FUNCTION "LKinCtrl_FwdFrame" : Void   // FC35005, SCL
TITLE = LKinCtrl_FwdFrame
{ S7_Optimized_Access := 'TRUE' }
AUTHOR : tech.team.motioncontrol@siemens.com
FAMILY : LKinCtrl
VERSION : 1.1
// Functionality: This function is calculating a forward frame transformation (-> In: Position in frame, Out: Position without frame)
// Support: tech.team.motioncontrol@siemens.com
// Note: Parameter comments are only available in language 'English (United States)'
   VAR_INPUT
      xIn : LReal;   // Input value x
      yIn : LReal;   // Input value y
      zIn : LReal;   // Input value z
      mode : Int;   // 0: Rotation + Translation, else: Rotation only
      frame : "LKinCtrl_typeFrame";   // Frame
   END_VAR
   VAR_OUTPUT
      xOut : LReal;   // Output value x
      yOut : LReal;   // Output value y
      zOut : LReal;   // Output value z
   END_VAR
   VAR_TEMP
      tempX1 : LReal;
      tempY1 : LReal;
      tempZ1 : LReal;
      tempX2 : LReal;
      tempY2 : LReal;
      tempZ2 : LReal;
      tempSin : LReal;
      tempCos : LReal;
   END_VAR
   // Ret_Val : Return value
   VAR CONSTANT
      DEGRAD : LReal := 0.0174532925199433;
   END_VAR
BEGIN
   //================================================================================
   // SIEMENS AG
   // (c)Copyright 2018 All Rights Reserved
   //--------------------------------------------------------------------------------
   // Library: LKinCtrl 
   // Tested with: S7-1516T-3 PN
   // Engineering: TIA Portal V15
   // Restrictions: -
   // Requirements: S7-1500/S7-1500T FW 2.5
   // Functionality: LKinCtrl_FwdFrame
   // This function is calculating a forward frame transformation
   //                (-> In: Position in frame, Out: Position without frame)
   // Support: tech.team.motioncontrol@siemens.com
   // Note: Parameter comments are only available in language 'English (United States)'
   //--------------------------------------------------------------------------------
   // Change log table:
   // Version  Date       Expert in charge Changes applied
   // 01.00.00 29.03.2018 SF               created
   // 01.01.00 03.09.2018 SF               bugfix
   //================================================================================

   REGION INPUT
     #tempX1 := #xIn;
     #tempY1 := #yIn;
     #tempZ1 := #zIn;
   END_REGION

   REGION ROTATION
     //first step: rotate c -> b -> a
     //----------------------------------------------------------------------------
     IF (#frame.c <> 0.0) THEN //x-rotation neccessary?
       #tempSin := SIN(#frame.c * #DEGRAD);
       #tempCos := COS(#frame.c * #DEGRAD);
       //rotate
       #tempX2 := #tempX1;
       #tempY2 := #tempY1 * #tempCos - #tempZ1 * #tempSin;
       #tempZ2 := #tempY1 * #tempSin + #tempZ1 * #tempCos;
       //store  
       #tempX1 := #tempX2;
       #tempY1 := #tempY2;
       #tempZ1 := #tempZ2;
     END_IF;

     IF (#frame.b <> 0.0) THEN //y-rotation neccessary?
       #tempSin := SIN(#frame.b * #DEGRAD);
       #tempCos := COS(#frame.b * #DEGRAD);
       //rotate
       #tempX2 := #tempX1 * #tempCos + #tempZ1 * #tempSin;
       #tempY2 := #tempY1;
       #tempZ2 := - #tempX1 * #tempSin + #tempZ1 * #tempCos;
       //store  
       #tempX1 := #tempX2;
       #tempY1 := #tempY2;
       #tempZ1 := #tempZ2;
     END_IF;

     IF (#frame.a <> 0.0) THEN //z-rotation neccessary?
       #tempSin := SIN(#frame.a * #DEGRAD);
       #tempCos := COS(#frame.a * #DEGRAD);
       //rotate
       #tempX2 := #tempX1 * #tempCos - #tempY1 * #tempSin;
       #tempY2 := #tempX1 * #tempSin + #tempY1 * #tempCos;
       #tempZ2 := #tempZ1;
       //store  
       #tempX1 := #tempX2;
       #tempY1 := #tempY2;
       #tempZ1 := #tempZ2;
     END_IF;
   END_REGION

   REGION TRANSLATION
     IF #mode = 0 THEN
       //second step: translation/ shifting X,Y,Z
       //-------------------------------------------------------------------------
       IF (#frame.x <> 0.0) THEN
         #tempX1 := #tempX1 + #frame.x;
       END_IF;
       IF (#frame.y <> 0.0) THEN
         #tempY1 := #tempY1 + #frame.y;
       END_IF;
       IF (#frame.z <> 0.0) THEN
         #tempZ1 := #tempZ1 + #frame.z;
       END_IF;
     END_IF;
   END_REGION

   REGION OUTPUT
     #xOut := #tempX1;
     #yOut := #tempY1;
     #zOut := #tempZ1;
   END_REGION
END_FUNCTION

FUNCTION "LKinCtrl_InvFrame" : Void   // FC35006, SCL
TITLE = LKinCtrl_InvFrame
{ S7_Optimized_Access := 'TRUE' }
AUTHOR : tech.team.motioncontrol@siemens.com
FAMILY : LKinCtrl
VERSION : 1.1
// Functionality: This function is calculating a inverse frame transformation (-> In: Position without frame, Out: Position in frame)
// Support: tech.team.motioncontrol@siemens.com
// Note: Parameter comments are only available in language 'English (United States)'
   VAR_INPUT
      xIn : LReal;   // Input value x
      yIn : LReal;   // Input value y
      zIn : LReal;   // Input value z
      mode : Int;   // 0: Rotation + Translation, else: Rotation only
      frame : "LKinCtrl_typeFrame";   // Frame
   END_VAR
   VAR_OUTPUT
      xOut : LReal;   // Output value x
      yOut : LReal;   // Output value y
      zOut : LReal;   // Output value z
   END_VAR
   VAR_TEMP
      tempX1 : LReal;
      tempY1 : LReal;
      tempZ1 : LReal;
      tempX2 : LReal;
      tempY2 : LReal;
      tempZ2 : LReal;
      tempSin : LReal;
      tempCos : LReal;
   END_VAR
   // Ret_Val : Return value
   VAR CONSTANT
      DEGRAD : LReal := 0.0174532925199433;
   END_VAR
BEGIN
   //================================================================================
   // SIEMENS AG
   // (c)Copyright 2018 All Rights Reserved
   //--------------------------------------------------------------------------------
   // Library: LKinCtrl
   // Tested with: S7-1516T-3 PN
   // Engineering: TIA Portal V15
   // Restrictions: -
   // Requirements: S7-1500/S7-1500T FW 2.5
   // Functionality: LKinCtrl_InvFrame
   // This function is calculating a inverse frame transformation
   //                (-> In: Position without frame, Out: Position in frame)
   // Support: tech.team.motioncontrol@siemens.com
   // Note: Parameter comments are only available in language 'English (United States)'
   //--------------------------------------------------------------------------------
   // Change log table:
   // Version  Date       Expert in charge Changes applied
   // 01.00.00 29.03.2018 SF               created
   // 01.01.00 03.09.2018 SF               bugfix
   //================================================================================

   REGION INPUT
     #tempX1 := #xIn;
     #tempY1 := #yIn;
     #tempZ1 := #zIn;
   END_REGION

   REGION TRANSLATION
     IF #mode = 0 THEN
       //first step: translation/ shifting X,Y,Z
       //-------------------------------------------------------------------------
       IF (#frame.x <> 0.0) THEN
         #tempX1 := #tempX1 - #frame.x;
       END_IF;
       IF (#frame.y <> 0.0) THEN
         #tempY1 := #tempY1 - #frame.y;
       END_IF;
       IF (#frame.z <> 0.0) THEN
         #tempZ1 := #tempZ1 - #frame.z;
       END_IF;
     END_IF;
   END_REGION

   REGION ROTATION
     //second step: rotate a -> b -> c
     //---------------------------------------------------------------------------
     IF (#frame.a <> 0.0) THEN //z-rotation neccessary?
       #tempSin := SIN(#frame.a * #DEGRAD);
       #tempCos := COS(#frame.a * #DEGRAD);
       //rotate
       #tempX2 := #tempX1 * #tempCos + #tempY1 * #tempSin;
       #tempY2 := - #tempX1 * #tempSin + #tempY1 * #tempCos;
       #tempZ2 := #tempZ1;
       //store  
       #tempX1 := #tempX2;
       #tempY1 := #tempY2;
       #tempZ1 := #tempZ2;
     END_IF;

     IF (#frame.b <> 0.0) THEN //y-rotation neccessary?
       #tempSin := SIN(#frame.b * #DEGRAD);
       #tempCos := COS(#frame.b * #DEGRAD);
       //rotate
       #tempX2 := #tempX1 * #tempCos - #tempZ1 * #tempSin;
       #tempY2 := #tempY1;
       #tempZ2 := #tempX1 * #tempSin + #tempZ1 * #tempCos;
       //store  
       #tempX1 := #tempX2;
       #tempY1 := #tempY2;
       #tempZ1 := #tempZ2;
     END_IF;

     IF (#frame.c <> 0.0) THEN //x-rotation neccessary?
       #tempSin := SIN(#frame.c * #DEGRAD);
       #tempCos := COS(#frame.c * #DEGRAD);
       //rotate
       #tempX2 := #tempX1;
       #tempY2 := #tempY1 * #tempCos + #tempZ1 * #tempSin;
       #tempZ2 := - #tempY1 * #tempSin + #tempZ1 * #tempCos;
       //store  
       #tempX1 := #tempX2;
       #tempY1 := #tempY2;
       #tempZ1 := #tempZ2;
     END_IF;
   END_REGION

   REGION OUTPUT
     #xOut := #tempX1;
     #yOut := #tempY1;
     #zOut := #tempZ1;
   END_REGION
END_FUNCTION

FUNCTION "LKinCtrl_FrameTrans" : Void   // FC35007, SCL
TITLE = LKinCtrl_FrameTrans
{ S7_Optimized_Access := 'TRUE' }
AUTHOR : tech.team.motioncontrol@siemens.com
FAMILY : LKinCtrl
VERSION : 2.0
// The FC calculates a given position transformed into or from another coordinate system depending on the actual / previous coordinate system of the cmd
   VAR_INPUT
      coordSystem : DInt;   // actual coordinate system
      coordSystemOld : DInt;   // previous coordinate system
      OCSFrames : Array[1..3] of "LKinCtrl_typeFrame";   // frame parameters read from TO_Kinematics
   END_VAR
   VAR_IN_OUT
      position : Array[1..4] of LReal;   // position to be transformed
   END_VAR
BEGIN
   //==========================================================================================
   // SIEMENS AG
   // (c)Copyright 2020 All Rights Reserved
   //------------------------------------------------------------------------------------------
   // Library: LKinCtrl
   // Tested with: S7-1517T-3 PN/DP
   // Engineering: TIA Portal V15
   // Restrictions: ---
   // Requirements: S7-1500T FW 2.5
   // Functionality: LKinCtrl_FrameTrans
   // The FC calculates a given position transformed into or from another coordinate system
   // depending on the actual / previous coordinate system of the cmd
   // 
   // Support: tech.team.motioncontrol@siemens.com
   // Note: Parameter comments are only available in language 'English (United States)'
   //------------------------------------------------------------------------------------------
   // Change log table:
   // Version    Date          Expert in charge    Changes applied
   // 01.00.00   16.04.2019    JR                  First release version v1.0
   // 02.00.00   14.04.2020    FR                  Use array of frames
   //===========================================================================================

   // Check if last CS differs from actual CS
   IF #coordSystem = #coordSystemOld THEN
     // No calculation needed --> Return
     RETURN;
   END_IF;

   // Calc new position
   // =================
   // Check if last CS was a OCS
   // YES: Transform position to WCS
   // NO: Do nothing --> Position is already in WCS
   IF (#coordSystemOld >= "CS_OCS1" AND #coordSystemOld <= "CS_OCS3") THEN
     // Get frame to WCS
     // foward frame transformation of lastPos to interprete position in WCS instead of OCS[1..3]
     "LKinCtrl_FwdFrame"(xIn := #position[1],
                         yIn := #position[2],
                         zIn := #position[3],
                         mode := 0,
                         frame := #OCSFrames[#coordSystemOld],
                         xOut => #position[1],
                         yOut => #position[2],
                         zOut => #position[3]);

     // Add "a" rotation to pos[4]
     // Rotation is needed because no change of orientation shall be done
     #position[4] := #position[4] + #OCSFrames[#coordSystemOld].a;
   ELSE
     ; // We are already in WCS
   END_IF;

   // Check if target CS is a OCS
   // YES: Transform position to target OCS
   // NO: Target CS is WCS --> Position is already in WCS from above
   IF (#coordSystem >= "CS_OCS1" AND #coordSystem <= "CS_OCS3") THEN
     // Get frame to target OCS
     // inverse frame transformation of lastPos to interprete position in OCS[1..3] instead of WCS
     "LKinCtrl_InvFrame"(xIn := #position[1],
                         yIn := #position[2],
                         zIn := #position[3],
                         mode := 0,
                         frame := #OCSFrames[#coordSystem],
                         xOut => #position[1],
                         yOut => #position[2],
                         zOut => #position[3]);

     // Substract "a" rotation to pos[4]
     // Rotation is needed because no change of orientation shall be done
     #position[4] := #position[4] - #OCSFrames[#coordSystem].a;
   ELSE
     ; // We are already in WCS
   END_IF;
END_FUNCTION

FUNCTION "LKinCtrl_ConvCircMode3To1" : Word   // FC35008, SCL
TITLE = LKinCtrl_ConvCircMode3To1
{ S7_Optimized_Access := 'TRUE' }
AUTHOR : tech.team.motioncontrol@siemens.com
FAMILY : LKinCtrl
VERSION : 2.0
// The FC converts a circular motion command programmed with circMode 3 (GCode) to a circular command programmed with circMode 1 (center point and arc given)
   VAR_INPUT
      coordinates : Variant;   // endPoint from path data element
      lastPos : Array[1..4] of LReal;   // previous last position
   END_VAR
   VAR_OUTPUT
      errorMessage : String;   // error message
   END_VAR
   VAR_IN_OUT
      cmdType : Int;   // cmdType of path data element
      circleParameters : "LKinCtrl_typeCircleParameters";   // circle parameters of path data element
   END_VAR
   VAR_TEMP
      tempAuxPoint : Array[1..3] of LReal;   // resulting auxPoint
      tempEndPointResult : Array[1..4] of LReal;   // resulting endPoint
      tempOM : Array[1..2] of LReal;   // temporary math variable
      tempMS : Array[1..2] of LReal;   // temporary math variable
      tempME : Array[1..2] of LReal;   // temporary math variable
      tempAxisVector : Array[1..2] of LReal;   // temporary math variable
      tempScalarProd_ME_Axis : LReal;   // temporary math variable
      tempScalarProd_MS_Axis : LReal;   // temporary math variable
      tempLength_ME : LReal;   // temporary math variable
      tempLength_MS : LReal;   // temporary math variable
      tempAngleME_rad : LReal;   // temporary math variable
      tempAngleMS_rad : LReal;   // temporary math variable
      tempAngleME_deg : LReal;   // temporary math variable
      tempAngleMS_deg : LReal;   // temporary math variable
      tempAngleDiff_deg : LReal;   // temporary math variable
      tempCtr : Int;   // temporary counter
      tempCoordinatesArray : REF_TO Array[1..4] of LReal;   // reference to coordinates from pre buf element
      tempCoordinatesStruct : REF_TO "LKinCtrl_typeCartesianPosition";   // reference to coordinates from normal element
      tempCoordinates : Array[1..4] of LReal;   // temporary array for input end point
   END_VAR
   // Ret_Val : return value
   VAR CONSTANT
      ERR_INVALID_CMDTYPE : Word := 16#8265;   // error due to invalid cmdType
      STATUS_NO_ERROR : Word := 16#0;   // status no error occured
   END_VAR
BEGIN
   //==========================================================================================
   // SIEMENS AG
   // (c)Copyright 2020 All Rights Reserved
   //------------------------------------------------------------------------------------------
   // Library: LKinCtrl
   // Tested with: S7-1517T-3 PN/DP
   // Engineering: TIA Portal V15
   // Restrictions: ---
   // Requirements: S7-1500T FW 2.5
   // Functionality: LKinCtrl_ConvCircMode3To1
   // The FC converts a circular motion command programmed with circMode 3 (GCode) to a circular
   // command programmed with circMode 1 (center point and arc given)
   // 
   // Support: tech.team.motioncontrol@siemens.com
   // Note: Parameter comments are only available in language 'English (United States)'
   //------------------------------------------------------------------------------------------
   // Change log table:
   // Version    Date          Expert in charge    Changes applied
   // 01.00.00   03.07.2019    JR                  First release version v1.0
   // 02.00.00   06.04.2020    FR                  Changed interface to fit PathDataPreBuf and normal element
   //===========================================================================================

   IF TypeOf(#coordinates) = LKinCtrl_typeCartesianPosition THEN
     // Assignment
     #tempCoordinatesStruct ?= #coordinates;

     // Assign temp with values
     #tempCoordinates[1] := #tempCoordinatesStruct<?OpDeref?>.x;
     #tempCoordinates[2] := #tempCoordinatesStruct<?OpDeref?>.y;
     #tempCoordinates[3] := #tempCoordinatesStruct<?OpDeref?>.z;
     #tempCoordinates[4] := #tempCoordinatesStruct<?OpDeref?>.a;

   ELSIF TypeOfElements(#coordinates) = LReal AND IS_ARRAY(#coordinates) AND CountOfElements(#coordinates) = 4 THEN
     // Assignment
     #tempCoordinatesArray ?= #coordinates;

     // Assign temp with values
     #tempCoordinates := #tempCoordinatesArray<?OpDeref?>;

   ELSE
     ; // Wrong input ?
   END_IF;

   // add conversion of circMode CM: 3 circular cmds -> CM: 1
   IF (#cmdType = "LKINCTRL_MC_MOVECIRCULARABS"
     OR #cmdType = "LKINCTRL_MC_MOVECIRCULARREL")
     AND #circleParameters.circMode = 3
   THEN

     // conversion relative to absoulte for auxPoint (and EndPoint)
     FOR #tempCtr := 1 TO 3 DO
       // always convert auxPoint ==> always relative in this circle definition
       // add new auxPoint as incremental value to last position
       #tempAuxPoint[#tempCtr] := #lastPos[#tempCtr] + #circleParameters.auxPoint[#tempCtr];
       // copy edited auxPoint to command for later use
       #circleParameters.auxPoint[#tempCtr] := #tempAuxPoint[#tempCtr];
     END_FOR;

     // only convert endPoint in case of relative command
     IF #cmdType = "LKINCTRL_MC_MOVECIRCULARREL" THEN
       #tempEndPointResult[1] := #lastPos[1] + #tempCoordinates[1];
       #tempEndPointResult[2] := #lastPos[2] + #tempCoordinates[2];
       #tempEndPointResult[3] := #lastPos[3] + #tempCoordinates[3];
       #tempEndPointResult[4] := #lastPos[4] + #tempCoordinates[4];
       #cmdType := "LKINCTRL_MC_MOVECIRCULARABS";
     ELSE
       #tempEndPointResult := #tempCoordinates;
     END_IF;

     // change circMode = 3 (define center and endPoint) to circMode = 1 (define center and arc)
     #circleParameters.circMode := 1;

     // different behavior for different circlePlanes - write input vectors to calc variables 2D
     // 0: ciclePlane XZ
     IF #circleParameters.circlePlane = 0 THEN

       // vector origin to circle center point 
       #tempOM[1] := #tempAuxPoint[1];
       #tempOM[2] := #tempAuxPoint[3];

       // unit vector x axis
       #tempAxisVector[1] := 1;
       #tempAxisVector[2] := 0;

       // vector circle center point to start point
       #tempMS[1] := #lastPos[1] - #tempOM[1];
       #tempMS[2] := #tempOM[2] - #lastPos[3];

       // vector circle center point to end point
       #tempME[1] := #tempEndPointResult[1] - #tempOM[1];
       #tempME[2] := #tempOM[2] - #tempEndPointResult[3];

       // 1: ciclePlane YZ
     ELSIF #circleParameters.circlePlane = 1 THEN

       // vector origin to circle center point 
       #tempOM[1] := #tempAuxPoint[2];
       #tempOM[2] := #tempAuxPoint[3];

       // unit vector x axis ==> simulating y axis here due to moved commands
       #tempAxisVector[1] := 1;
       #tempAxisVector[2] := 0;

       // vector circle center point to start point
       #tempMS[1] := #lastPos[2] - #tempOM[1];
       #tempMS[2] := #lastPos[3] - #tempOM[2];

       // vector circle center point to end point
       #tempME[1] := #tempEndPointResult[2] - #tempOM[1];
       #tempME[2] := #tempEndPointResult[3] - #tempOM[2];

       // 2: ciclePlane XY
     ELSIF #circleParameters.circlePlane = 2 THEN

       // vector origin to circle center point 
       #tempOM[1] := #tempAuxPoint[1];
       #tempOM[2] := #tempAuxPoint[2];

       // unit vector x axis
       #tempAxisVector[1] := 1;
       #tempAxisVector[2] := 0;


       // vector circle center point to start point
       #tempMS[1] := #lastPos[1] - #tempOM[1];
       #tempMS[2] := #lastPos[2] - #tempOM[2];

       // vector circle center point to end point
       #tempME[1] := #tempEndPointResult[1] - #tempOM[1];
       #tempME[2] := #tempEndPointResult[2] - #tempOM[2];

     ELSE
       // error ==> wrong circlePlane
       ;
     END_IF;

     // VECTOR CALCULATIONS
     // calc scalar product of ME (circle center point to end point) with x axis
     #tempScalarProd_ME_Axis := "LKinCtrl_VecScalarProd_2D"(vIn1 := #tempME, vIn2 := #tempAxisVector);
     // calc scalar product of MS (circle center point to start point / LastPos) with x axis
     #tempScalarProd_MS_Axis := "LKinCtrl_VecScalarProd_2D"(vIn1 := #tempMS, vIn2 := #tempAxisVector);

     // calc vector length ME
     #tempLength_ME := "LKinCtrl_VecAbs_2D"(#tempME);
     // calc vector length MS
     #tempLength_MS := "LKinCtrl_VecAbs_2D"(#tempMS);

     // calc angle ME to axis
     #tempAngleME_rad := ACOS(#tempScalarProd_ME_Axis / (#tempLength_ME * 1));

     IF #tempME[2] <= 0 THEN
       // invert angle due to ACOS range (only 0..PI)
       #tempAngleME_rad := 2 * "LKINCTRL_PI" - #tempAngleME_rad;
     ELSE
       ;
     END_IF;
     // convert to degrees
     #tempAngleME_deg := #tempAngleME_rad * 180 / "LKINCTRL_PI";

     // calc angle MS to axis
     #tempAngleMS_rad := ACOS(#tempScalarProd_MS_Axis / (#tempLength_MS * 1));
     // check for vector Ms to point downwards (below ! (x) axis)
     IF #tempMS[2] < 0 THEN
       // invert angle due to ACOS range
       #tempAngleMS_rad := 2 * "LKINCTRL_PI" - #tempAngleMS_rad;
     ELSE
       ;
     END_IF;
     // convert to degrees
     #tempAngleMS_deg := #tempAngleMS_rad * 180 / "LKINCTRL_PI";


     // separation of path choice for angle calculation
     // 0: CCW - counterclockwise / mathematical positive angle
     IF #circleParameters.pathChoice = 0 THEN
       // calculate difference angle
       #tempAngleDiff_deg := #tempAngleME_deg - #tempAngleMS_deg;
       IF #tempAngleDiff_deg > 0 THEN
         // write caclulated angle
         #circleParameters.arc := #tempAngleDiff_deg;
       ELSE
         // write caclulated angle ==> add 360 degrees to get positive angle value
         #circleParameters.arc := #tempAngleDiff_deg + 360;
       END_IF;

       // 1: CW - clockwise / mathematical negative angle
     ELSIF #circleParameters.pathChoice = 1 THEN
       // calculate difference angle
       #tempAngleDiff_deg := #tempAngleMS_deg - #tempAngleME_deg;
       IF #tempAngleDiff_deg >(* = *) 0 THEN
         // write caclulated angle
         #circleParameters.arc := #tempAngleDiff_deg;
       ELSE
         // write caclulated angle ==> add 360 degrees to get positive angle value
         #circleParameters.arc := #tempAngleDiff_deg + 360;
       END_IF;

     ELSE
       // wrong input for pathChoice
       ;
     END_IF;
     // conversion successful
     #LKinCtrl_ConvCircMode3To1 := #STATUS_NO_ERROR;

   ELSE
     // do nothing
     #LKinCtrl_ConvCircMode3To1 := #ERR_INVALID_CMDTYPE;
     #errorMessage := 'no circular command to convert';
   END_IF;
END_FUNCTION

FUNCTION "LKinCtrl_EvaluateParamValidBits" : Void   // FC35009, SCL
TITLE = LKinCtrl_EvaluateParamValidBits
{ S7_Optimized_Access := 'TRUE' }
AUTHOR : tech.team.motioncontrol@siemens.com
FAMILY : LKinCtrl
VERSION : 1.0
// The FC evaluates the parameterValid bits of a given command and copies the coordinates for valid bits and overwrites coordinates by last position or 0.0 increment for invalid bits.
   VAR_INPUT
      parameterValidBits : Array[1.."LKINCTRL_NO_OF_VALID_BITS"] of Bool;   // parameter valid bits of actual command
      lastPos : Array[1..4] of LReal;   // previous last position
   END_VAR
   VAR_OUTPUT
      errorMessage : String;   // error message
   END_VAR
   VAR_IN_OUT
      command : "LKinCtrl_typePathDataElement";   // command to evaluate and edit
   END_VAR
   VAR_TEMP
      tempPosElemCtr : Int;   // temporary counter variable
   END_VAR
BEGIN
   //==========================================================================================
   // SIEMENS AG
   // (c)Copyright 2019 All Rights Reserved
   //------------------------------------------------------------------------------------------
   // Library: LKinCtrl
   // Tested with: S7-1517T-3 PN/DP
   // Engineering: TIA Portal V15
   // Restrictions: ---
   // Requirements: S7-1500T FW 2.5
   // Functionality: LKinCtrl_EvaluateParamValidBits
   // The FC evaluates the parameterValid bits of a given command and copies the coordinates for
   // valid bits and overwrites coordinates by last position or 0.0 increment for invalid bits.
   // 
   // Support: tech.team.motioncontrol@siemens.com
   // Note: Parameter comments are only available in language 'English (United States)'
   //------------------------------------------------------------------------------------------
   // Change log table:
   // Version    Date          Expert in charge    Changes applied
   // 01.00.00   08.07.2019    JR                  First release version v1.0
   // 01.00.01   09.08.2019    JR                  excluded auxPoint from parameter valid bits
   //===========================================================================================

   // ParameterValid bit check
   //====================================================================================================================================

   // -----------------------------------------------------------------------------------
   IF #command.cmdType = "LKINCTRL_MC_MOVELINEARABS" OR #command.cmdType = "LKINCTRL_MC_MOVECIRCULARABS" THEN

     FOR #tempPosElemCtr := 1 TO "LKINCTRL_NO_OF_VALID_BITS" DO
       // Check valid bits and copy last pos (X,Y,Z,A) where missing
       IF #parameterValidBits[#tempPosElemCtr] = FALSE THEN
         // write lastPos as target pos if invalid
         IF #tempPosElemCtr = 1 THEN
           #command.cmdCoordinates.cartesianPosition.x := #lastPos[#tempPosElemCtr];
         ELSIF #tempPosElemCtr = 2 THEN
           #command.cmdCoordinates.cartesianPosition.y := #lastPos[#tempPosElemCtr];
         ELSIF #tempPosElemCtr = 3 THEN
           #command.cmdCoordinates.cartesianPosition.z := #lastPos[#tempPosElemCtr];
         ELSIF #tempPosElemCtr = 4 THEN
           #command.cmdCoordinates.cartesianPosition.a := #lastPos[#tempPosElemCtr];
         END_IF;

         // // exclude auxPoint from parameterValidBits, add additional parameterValidBits if needed
         // // write lastPos to auxPoint if invalid
         // IF #tempPosElemCtr < 4 THEN
         //   #command.cmdParameters.circleParameters.auxPoint[#tempPosElemCtr] := #lastPos[#tempPosElemCtr];
         // ELSE
         //   ; // do not copy for tempPosElemCtr = 4
         // END_IF;
       ELSE
         ; // Keep programmed position from #pathDataElementPreBuf.cmdCoordinates.cartesianPosition
       END_IF;
     END_FOR;

   ELSIF #command.cmdType = "LKINCTRL_MC_MOVELINEARREL" OR #command.cmdType = "LKINCTRL_MC_MOVECIRCULARREL" THEN
     FOR #tempPosElemCtr := 1 TO "LKINCTRL_NO_OF_VALID_BITS" DO
       // Check valid bits and set absolute pos to 0.0 (X,Y,Z,A)
       IF #parameterValidBits[#tempPosElemCtr] = FALSE THEN
         // write no increment as relative target pos if invalid
         IF #tempPosElemCtr = 1 THEN
           #command.cmdCoordinates.cartesianPosition.x := 0.0;
         ELSIF #tempPosElemCtr = 2 THEN
           #command.cmdCoordinates.cartesianPosition.y := 0.0;
         ELSIF #tempPosElemCtr = 3 THEN
           #command.cmdCoordinates.cartesianPosition.z := 0.0;
         ELSIF #tempPosElemCtr = 4 THEN
           #command.cmdCoordinates.cartesianPosition.a := 0.0;
         END_IF;

         // // exclude auxPoint from parameterValidBits, add additional parameterValidBits if needed
         // // write no increment as relative target pos if invalid
         // IF #tempPosElemCtr < 4 THEN
         //   #command.cmdParameters.circleParameters.auxPoint[#tempPosElemCtr] := 0.0;
         // ELSE
         //   ; // do not copy for tempPosElemCtr = 4
         // END_IF;
       ELSE
         ; // Keep programmed position from #pathDataElementPreBuf.cmdCoordinates.cartesianPosition
       END_IF;
     END_FOR;
   ELSE
     ; // Nothing to do for this cmdType
   END_IF;
END_FUNCTION

FUNCTION "LKinCtrl_CallMC_TrackConv_PosAxis" : Void   // FC35010, SCL
TITLE = LKinCtrl_CallMC_TrackConv_PosAxis
{ S7_Optimized_Access := 'TRUE' }
AUTHOR : tech.team.motioncontrol@siemens.com
FAMILY : LKinCtrl
VERSION : 1.0
// Call given MC_TrackConveyorBelt instance
   VAR_INPUT
      posAxis : TO_PositioningAxis;   // Positioning axis input
      axesGroup : TO_Kinematics;   // Kinematics input
   END_VAR
   VAR_IN_OUT
      instTrackConveyorBelt : MC_TRACKCONVEYORBELT;   // Instance of MC_TrackConveyorBelt to be called
   END_VAR
BEGIN
   //================================================================================
   // SIEMENS AG
   // (c)Copyright 2020 All Rights Reserved
   //--------------------------------------------------------------------------------
   // Library: LKinCtrl
   // Tested with: S7-1517T-3 PN
   // Engineering: TIA Portal V16
   // Restrictions: -
   // Requirements: S7-1500T FW 2.8
   // Functionality: Call MC_TrackConveyorBelt
   // Support: tech.team.motioncontrol@siemens.com
   // Note: Parameter comments are only available in language 'English (United States)'
   //-----------------------------------------------------------------------------
   // Change log table:
   // Version    Date          Expert in charge    Changes applied
   // 01.00.00   24.04.2020    FR                  First released version
   //===========================================================================================

   // call MC_TrackConveyorBelt
   #instTrackConveyorBelt(AxesGroup:=#axesGroup,
                              ConveyorBelt:=#posAxis);
END_FUNCTION

FUNCTION "LKinCtrl_CallMC_TrackConv_SyncAxis" : Void   // FC35011, SCL
TITLE = LKinCtrl_CallMC_TrackConv_SyncAxis
{ S7_Optimized_Access := 'TRUE' }
AUTHOR : tech.team.motioncontrol@siemens.com
FAMILY : LKinCtrl
VERSION : 1.0
// Call given MC_TrackConveyorBelt instance
   VAR_INPUT
      syncAxis : TO_SynchronousAxis;   // Synchronous axis input
      axesGroup : TO_Kinematics;   // Kinematics input
   END_VAR
   VAR_IN_OUT
      instTrackConveyorBelt : MC_TRACKCONVEYORBELT;   // Instance of MC_TrackConveyorBelt to be called
   END_VAR
BEGIN
   //================================================================================
   // SIEMENS AG
   // (c)Copyright 2020 All Rights Reserved
   //--------------------------------------------------------------------------------
   // Library: LKinCtrl
   // Tested with: S7-1517T-3 PN
   // Engineering: TIA Portal V16
   // Restrictions: -
   // Requirements: S7-1500T FW 2.8
   // Functionality: Call MC_TrackConveyorBelt
   // Support: tech.team.motioncontrol@siemens.com
   // Note: Parameter comments are only available in language 'English (United States)'
   //-----------------------------------------------------------------------------
   // Change log table:
   // Version    Date          Expert in charge    Changes applied
   // 01.00.00   24.04.2020    FR                  First released version
   //===========================================================================================

   // call MC_TrackConveyorBelt
   #instTrackConveyorBelt(AxesGroup := #axesGroup,
                          ConveyorBelt := #syncAxis);
END_FUNCTION

FUNCTION "LKinCtrl_CallMC_TrackConv_ExtEncoder" : Void   // FC35012, SCL
TITLE = LKinCtrl_CallMC_TrackConv_ExtEncoder
{ S7_Optimized_Access := 'TRUE' }
AUTHOR : tech.team.motioncontrol@siemens.com
FAMILY : LKinCtrl
VERSION : 1.0
// Call given MC_TrackConveyorBelt instance
   VAR_INPUT
      extEncoder : TO_ExternalEncoder;   // External Encoder input
      axesGroup : TO_Kinematics;   // Kinematics input
   END_VAR
   VAR_IN_OUT
      instTrackConveyorBelt : MC_TRACKCONVEYORBELT;   // Instance of MC_TrackConveyorBelt to be called
   END_VAR
BEGIN
   //================================================================================
   // SIEMENS AG
   // (c)Copyright 2020 All Rights Reserved
   //--------------------------------------------------------------------------------
   // Library: LKinCtrl
   // Tested with: S7-1517T-3 PN
   // Engineering: TIA Portal V16
   // Restrictions: -
   // Requirements: S7-1500T FW 2.8
   // Functionality: Call MC_TrackConveyorBelt
   // Support: tech.team.motioncontrol@siemens.com
   // Note: Parameter comments are only available in language 'English (United States)'
   //-----------------------------------------------------------------------------
   // Change log table:
   // Version    Date          Expert in charge    Changes applied
   // 01.00.00   24.04.2020    FR                  First released version
   //===========================================================================================

   // call MC_TrackConveyorBelt
   #instTrackConveyorBelt(AxesGroup := #axesGroup,
                          ConveyorBelt := #extEncoder);
END_FUNCTION

FUNCTION "LKinCtrl_CallMC_TrackConv_LeadingAxisProxy" : Void   // FC35013, SCL
TITLE = LKinCtrl_CallMC_TrackConv_LeadingAxisProxy
{ S7_Optimized_Access := 'TRUE' }
AUTHOR : tech.team.motioncontrol@siemens.com
FAMILY : LKinCtrl
VERSION : 1.0
// Call given MC_TrackConveyorBelt instance
   VAR_INPUT
      leadingAxisProxy : TO_LeadingAxisProxy;   // Leading axis proxy input
      axesGroup : TO_Kinematics;   // Kinematics input
   END_VAR
   VAR_IN_OUT
      instTrackConveyorBelt : MC_TRACKCONVEYORBELT;   // Instance of MC_TrackConveyorBelt to be called
   END_VAR
BEGIN
   //================================================================================
   // SIEMENS AG
   // (c)Copyright 2020 All Rights Reserved
   //--------------------------------------------------------------------------------
   // Library: LKinCtrl
   // Tested with: S7-1517T-3 PN
   // Engineering: TIA Portal V16
   // Restrictions: -
   // Requirements: S7-1500T FW 2.8
   // Functionality: Call MC_TrackConveyorBelt
   // Support: tech.team.motioncontrol@siemens.com
   // Note: Parameter comments are only available in language 'English (United States)'
   //-----------------------------------------------------------------------------
   // Change log table:
   // Version    Date          Expert in charge    Changes applied
   // 01.00.00   24.04.2020    FR                  First released version
   //===========================================================================================

   // call MC_TrackConveyorBelt
   #instTrackConveyorBelt(AxesGroup := #axesGroup,
                          ConveyorBelt := #leadingAxisProxy);
END_FUNCTION

FUNCTION "LKinCtrl_VecAbs_2D" : LReal   // FC35029, SCL
TITLE = LKinCtrl_VecAbs_2D
{ S7_Optimized_Access := 'TRUE' }
AUTHOR : tech.team.motioncontrol@siemens.com
FAMILY : LKinCtrl
VERSION : 1.0
// Calculates the length of a given vector in 2D
   VAR_INPUT
      vIn : Array[1..2] of LReal;   // Input vector
   END_VAR
   // Ret_Val : Output scalar
BEGIN
   //=============================================================================
   // SIEMENS AG
   // (c)Copyright 2019 All Rights Reserved
   //-----------------------------------------------------------------------------
   // Library: - 
   // Tested with: S7-1516T-3 PN
   // Engineering: TIA Portal V15
   // Restrictions: -
   // Requirements: S7-1500/S7-1500T FW 2.5
   // Functionality: Calculate length of vector
   //-----------------------------------------------------------------------------
   // Change log table:
   // Version  Date       Expert in charge Changes applied
   // 01.00.00 27.08.2018 SF               created
   // 01.00.01 29.01.2019 JR               adaptions for LKinCtrl 
   //=============================================================================

   #LKinCtrl_VecAbs_2D := SQRT((* #vIn[0]*#vIn[0] + *)#vIn[1]*#vIn[1] + #vIn[2]*#vIn[2]);
END_FUNCTION

FUNCTION "LKinCtrl_VecScalarProd_2D" : LReal   // FC35030, SCL
TITLE = LKinCtrl_VecScalarProd_2D / LKinCtrl_VecScalarProd
{ S7_Optimized_Access := 'TRUE' }
AUTHOR : tech.team.motioncontrol@siemens.com
FAMILY : LKinCtrl
VERSION : 1.0
// Calculates the scalar product of given vectors
   VAR_INPUT
      vIn1 : Array[1..2] of LReal;   // Input vector 1
      vIn2 : Array[1..2] of LReal;   // Input vector 2
   END_VAR
   // Ret_Val : Output scalar
BEGIN
   //=============================================================================
   // SIEMENS AG
   // (c)Copyright 2019 All Rights Reserved
   //-----------------------------------------------------------------------------
   // Library: - 
   // Tested with: S7-1516T-3 PN
   // Engineering: TIA Portal V15
   // Restrictions: -
   // Requirements: S7-1500/S7-1500T FW 2.5
   // Functionality: Scalar product of two coordinates
   //-----------------------------------------------------------------------------
   // Change log table:
   // Version  Date       Expert in charge Changes applied
   // 01.00.00 27.08.2018 SF               created
   // 01.00.01 29.01.2019 JR               adaptions for LKinCtrl 
   //=============================================================================

   #LKinCtrl_VecScalarProd_2D := (* #vIn1[0]*#vIn2[0] + *)#vIn1[1]*#vIn2[1] + #vIn1[2]*#vIn2[2];
END_FUNCTION

FUNCTION "LKinCtrl_GetPathDataCmd" : Word   // FC35031, SCL
TITLE = LKinCtrl_GetPathDataCmd
{ S7_Optimized_Access := 'TRUE' }
AUTHOR : tech.team.motioncontrol@siemens.com
FAMILY : LKinCtrl
VERSION : 1.0
// Copy the path command from any path data type at the given index
   VAR_INPUT
      pathDataType : USInt;   // Type of path data which is connected
      index : DInt;   // Index to be copied
      pathDataReduced : REF_TO "LKinCtrl_typePathData_reduced";   // Reference to reduced path data
      pathData : REF_TO "LKinCtrl_typePathData";   // Reference to normal path data
      pathDataAdvanced : REF_TO "LKinCtrl_typePathData_advanced";   // Reference to advanced path data
   END_VAR
   VAR_OUTPUT
      pathDataCommand : "LKinCtrl_typePathDataElement";   // Resulting path data command
      parameterValid : Array[1.."LKINCTRL_NO_OF_VALID_BITS"] of Bool;   // Resulting parameter valid bits
   END_VAR
   VAR_TEMP
      tempCtr : Int;   // Temporary counter
   END_VAR
   // Ret_Val : Return value
BEGIN
   //==========================================================================================
   // SIEMENS AG
   // (c)Copyright 2020 All Rights Reserved
   //------------------------------------------------------------------------------------------
   // Library: LKinCtrl
   // Tested with: S7-1517T-3 PN/DP
   // Engineering: TIA Portal V15
   // Restrictions: ---
   // Requirements: S7-1500T FW 2.5
   // Functionality: LKinCtrl_GetPathDataCmd
   // The FC copies the path data command at the given index to the output.
   // 
   // Support: tech.team.motioncontrol@siemens.com
   // Note: Parameter comments are only available in language 'English (United States)'
   //------------------------------------------------------------------------------------------
   // Change log table:
   // Version    Date          Expert in charge    Changes applied
   // 01.00.00   07.04.2020    FR                  First release version v1.0
   //===========================================================================================

   // Set return value
   #LKinCtrl_GetPathDataCmd := 16#00;

   // Copy actual path data element where index is pointing at
   IF #pathDataType = "LKINCTRL_PATHDATA_TYPE_REDUCED" THEN
     // Copy command
     #pathDataCommand.cmdType := #pathDataReduced<?OpDeref?>.commands[#index].cmdType;
     #pathDataCommand.cmdName := #pathDataReduced<?OpDeref?>.commands[#index].cmdName;
     #pathDataCommand.cmdActivated := #pathDataReduced<?OpDeref?>.commands[#index].cmdActivated; // !
     #pathDataCommand.cmdCoordinates := #pathDataReduced<?OpDeref?>.commands[#index].cmdCoordinates;
     #pathDataCommand.cmdParameters.pathDynamics := #pathDataReduced<?OpDeref?>.commands[#index].cmdParameters.pathDynamics;
     #pathDataCommand.cmdParameters.orientationDirection := #pathDataReduced<?OpDeref?>.commands[#index].cmdParameters.orientationDirection;
     #pathDataCommand.cmdParameters.bufferMode := #pathDataReduced<?OpDeref?>.commands[#index].cmdParameters.bufferMode;
     #pathDataCommand.cmdParameters.transitionParameters := #pathDataReduced<?OpDeref?>.commands[#index].cmdParameters.transitionParameters;
     #pathDataCommand.cmdParameters.dynamicAdaption := #pathDataReduced<?OpDeref?>.commands[#index].cmdParameters.dynamicAdaption;
     #pathDataCommand.setFlags := #pathDataReduced<?OpDeref?>.commands[#index].setFlags;
     #pathDataCommand.valueFlags := #pathDataReduced<?OpDeref?>.commands[#index].valueFlags;

     // always set valid bits to true
     FOR #tempCtr := 1 TO "LKINCTRL_NO_OF_VALID_BITS" DO
       // Statement section FOR
       #parameterValid[#tempCtr] := TRUE;
     END_FOR;

   ELSIF #pathDataType = "LKINCTRL_PATHDATA_TYPE_NORMAL" THEN
     // Copy command
     #pathDataCommand := #pathData<?OpDeref?>.commands[#index];

     // always set valid bits to true
     FOR #tempCtr := 1 TO "LKINCTRL_NO_OF_VALID_BITS" DO
       // Statement section FOR
       #parameterValid[#tempCtr] := TRUE;
     END_FOR;

   ELSIF #pathDataType = "LKINCTRL_PATHDATA_TYPE_ADVANCED" THEN
     // Copy command
     #pathDataCommand.cmdType := #pathDataAdvanced<?OpDeref?>.commands[#index].cmdType;
     #pathDataCommand.cmdName := #pathDataAdvanced<?OpDeref?>.commands[#index].cmdName;
     #pathDataCommand.cmdActivated := #pathDataAdvanced<?OpDeref?>.commands[#index].cmdActivated;
     #pathDataCommand.cmdCoordinates := #pathDataAdvanced<?OpDeref?>.commands[#index].cmdCoordinates;
     #pathDataCommand.cmdParameters := #pathDataAdvanced<?OpDeref?>.commands[#index].cmdParameters;
     #pathDataCommand.setFlags := #pathDataAdvanced<?OpDeref?>.commands[#index].setFlags;
     #pathDataCommand.valueFlags := #pathDataAdvanced<?OpDeref?>.commands[#index].valueFlags;

     // Copy valid bits from command
     #parameterValid := #pathDataAdvanced<?OpDeref?>.commands[#index].parameterValid;

   ELSE
     // Set return value to error
     #LKinCtrl_GetPathDataCmd := 16#01;
   END_IF;
END_FUNCTION

// folder: LKinLang_Blocks

FUNCTION_BLOCK "LKinLang_Parser"   // FB35450, SCL
TITLE = LKinLang_Parser
{ S7_Optimized_Access := 'TRUE' }
AUTHOR : tech.team.motioncontrol@siemens.com
FAMILY : LKinLang
VERSION : 1.3
// The FB parses strings from line buffer to PathData commands using different language
// packages.
// The FB parses strings from line buffer to PathData commands using different languagepackages.
   VAR_INPUT
      execute : Bool;   // Rising edge starts action once
      stop : Bool;   // Rising edge stops execution
      language : Int;   // Selected language to be parsed
      syntaxCheck : USInt;   // 0: No check before; 1: Check only; 2: Check and execute
      flagModeDefaults : "LKinLang_typeFlagModeDefaults";   // Structure to define default flag settings for setFlags and valueFlags
   END_VAR
   VAR_OUTPUT
      done : Bool;   // TRUE: Commanded functionality has been completed successfully
      busy : Bool;   // TRUE: FB is not finished and new output values can be expected
      commandAborted : Bool;   // TRUE: Commanded functionality has been aborted by another command
      error : Bool;   // TRUE: An error occurred during the execution of the FB
      status : Word := 16#7000;   // 16#0000 - 16#7FFF: Status of the FB, 16#8000 - 16#FFFF: Error identification
      errorString : String;   // Error description as string
   END_VAR
   VAR_IN_OUT
      lineBuffer : "LKinLang_typeLineBuffer";   // String buffer connection
      pathData : "LKinCtrl_typePathData_advanced";   // PathData connection
      preProcessConfig : "LKinLang_typePreProcessorReplacement";   // Array which defines replacements
      parameterDefaults : Variant;   // Structure to define default values in language (e.g. velocity for rapid linear)
      interfaceVariables : "LKinLang_typeInterfaceVariables";   // Interface variables arrays
   END_VAR
   VAR
      statExecuteOld : Bool;   // Old value of 'execute' input for edge detection
      statDone : Bool;   // Static value for output 'done'
      statBusy : Bool;   // Static value for output 'busy'
      statCommandAborted : Bool;   // Static value for output 'commandAborted'
      statError : Bool;   // Static value for output 'error'
      statStatus : Word := 16#7000;   // Static value for output 'status'
      statErrorString : String;   // Error string variable
      statStopOld : Bool;   // Static storing for the stop input
      statFBState : DInt := 0;   // State in the state machine of the FB
      statStateIntern : Int;   // Internal state variable
      statSelectedLanguage : Int;   // Selected Language
      statPositioningMode : Int := 1;   // Positioning mode: 1=Absolute, 2=Relative
      statPositioningModeOld : Int := 1;   // Last Positioning mode
      statLastIndexLookUp : DInt;   // Last found command in Language Package
      statLastIndexOfMerger : Int;   // Last entry in merger array
      statLookUpTableCounter : Int;   // Counter to continue look up table
      statAddPointer : Int;   // Internal static to for the PathData add pointer
      statActualValueFlagNumber : Int;   // Static storing for the actual value flag number
      statActualFlagNumber : Int;   // Static storing for the actual boolean flag number
      statStringExpression : String;   // Static storing for the string expression
      statRightSideOfEquation : Bool;   // Static storing if right side of equation
      statDirectCmdWord : Word;   // Static storing direct command word
      statSyntaxCheck : USInt;   // Static storing for syntaxCheck input
      statSearchedLine : UDInt;   // Static storing for requested line number
      statConfigCmdWords : Array[1.."LKINLANG_NUMBER_OF_FOLLOW_VALUES"] of Word;   // Static storing config command word
      statTokenCheck : Struct   // Static struct with the token to check
         actual : String;
         previous : String;
      END_STRUCT;
      statTokenizedLine : "LKinLang_typeLineTokens";   // Tokenized line (String into separate strings)
      statSeparators : Array[1.."LKINLANG_NUMBER_OF_SEPARATORS"] of Byte;   // Array to save separators
      statMergers : Array[1.."LKINLANG_NUMBER_OF_MERGERS"] of Byte;   // Array to save mergers
      statActualCommand : "LKinLang_typePathDataElement";   // Path data command
      statActualCommandOld : "LKinLang_typePathDataElement";   // Last path data command
      statModalCommand : "LKinLang_typePathDataElement";   // Command Modal values
      statModalCommandOld : "LKinLang_typePathDataElement";   // Last command modal values
      statModalProgram : "LKinLang_typePathDataElement";   // Program modal values
      statPathDataElementEmpty : "LKinLang_typePathDataElement";   // Delete Path Data element
      statSetParametersInLine : Array[1.."LKINLANG_NUMBER_OF_CONDITIONS"] of "LKinLang_typeCondition";   // Conditions which were set in Line
      statSetParametersInCmd : Array[1.."LKINLANG_NUMBER_OF_CONDITIONS"] of "LKinLang_typeCondition";   // Conditions which were set in Cmd
      statSetParametersInPrg : Array[1.."LKINLANG_NUMBER_OF_CONDITIONS"] of "LKinLang_typeCondition";   // Conditions which were set in Prg
      statConditionsToCheck : Array[1.."LKINLANG_NUMBER_OF_CONDITIONS"] of "LKinLang_typeCondition";   // Conditions which have to be checked
      statConditionEmpty : "LKinLang_typeCondition";   // Delete conditions
      statParameterLookUpTable : Array[1.."LKINLANG_MAX_NUMBER_OF_PARAMETERS"] of "LKinLang_typeParameterLookUp";   // Array to save parameters
      statElementCounter : "LKinLang_typePathDataElementCounter";   // Counter of cmd modal values
      statElementCounterInLine : "LKinLang_typePathDataElementCounter";   // Counter of element in one line
      statValidCounts : "LKinLang_typePathDataElementCounter";   // Array which defines how often a parameter can be set
      statElementCounterEmpty : "LKinLang_typePathDataElementCounter";   // Delete counter
      statParameterDefinition : "LKinLang_typeParameterDefinition";   // Static storing for parameter definition
      statParameterDefinitionEmpty : "LKinLang_typeParameterDefinition";   // Delete parameter definition
      statParameterValid : "LKinLang_typePathDataValid";   // Static storing if a parameter is valid
      statParameterValidEmpty : "LKinLang_typePathDataValid";   // Delete parameter valid
      statPathDataValue : "LKinLang_typeDiffElementaryDatatypes";   // Static storing for path data element values
      statModalCmdValue : "LKinLang_typeDiffElementaryDatatypes";   // Static storing for path data element command modal values
      statModalPrgValue : "LKinLang_typeDiffElementaryDatatypes";   // Static storing for path data element program modal values
      statKeyToken : "LKinLang_typeKeyToken";   // Static storing different keywords
      statVariableDeclaration : "LKinLang_typeVariableDeclaration";   // Static storing the definition string for local and global variables
      statGlobalVariableDefinition : "LKinLang_typeLocalVarDefinition";   // Static storing the tokenized definition for global variables
      statLocalVariableDefinition : "LKinLang_typeLocalVarDefinition";   // Static storing the tokenized definition for local variables / Static storing the definition string for local variables
      statVariables : "LKinLang_typeLocalVariables";   // Structure containing local and global variables / Structure containing all local variables